FUNCTION "FC1041_TT_Taktimpuls" : Void   // FC1041, STL
TITLE = Taktimpuls bilden
{ S7_Optimized_Access := 'FALSE' }
AUTHOR : KT242
VERSION : 0.1
   VAR_INPUT
      IN_Drehfreigabe : Bool;   // Allgemeine Freigabe zum ansteuern der Anlage
      IN_Taktfreigabe : Bool;   // Freigabe zum Weitertakten der Anlage
      IN_Anlage_in_Position : Bool;   // Die Anlage befindet sich in der vorgegebenen Position
      IN_Start_Anlagenbetrieb : Bool;   // Die Anlage befindet sich in der Vorbereitung zum Produktionsbetrieb
      IN_Anlagenbetrieb : Bool;   // Die Anlage befindet sich im Produktionsbetrieb
      IN_DW_Taktzeit : S5Time;   // Zeitwert für die Taktzeit (Lauf- und Pausenzeit) der Anlage
      IN_Takttimer : Timer;   // Timer für die Bildung des Taktimpulses
      IN_Vorwarnzeit_1_in_Dec : Int;   // Zeitwert in Sekunden für eine Anfahrwarnung 1 vor dem Weitertakten
      IN_Vorwarnzeit_2_in_Dec : Int;   // Zeitwert in Sekunden für eine Anfahrwarnung 2 vor dem Weitertakten
   END_VAR
   VAR_IN_OUT
      IO_Status : "UDT_RT_Takt";   // Speichern der Takt- Zustände für das Programm
   END_VAR
   VAR_TEMP
      Temp_Restzeit : Int;   // Hilfwort mit Restzeit der Taktzeit in Sekunden
      Temp_Zeitraster : Byte;   // Hilfsbyte für dei ermittlung des Zeitrasters für die Bildung der Vorwarnungen
   END_VAR
BEGIN

REGION Network 1: Baustein abloeschen, wenn nicht Automatik
         O     #IN_Anlagenbetrieb;
         O     #IN_Start_Anlagenbetrieb;
         JC    NW1e;
   //
         R     #IO_Status.Vorwarnung_1;
         R     #IO_Status.Vorwarnung_2;
         R     #IO_Status.Taktzeit_beendet;
         R     #IO_Status.Taktimpuls;
         CLR;
         L     S5T#0MS;
         SP    #IN_Takttimer;
         BE;
   //
   NW1e: NOP   0;
END_REGION

REGION Network 2: Taktimpuls bilden
         L     #IN_DW_Taktzeit;
         A     #IN_Taktfreigabe;
         A     #IN_Drehfreigabe;
         A     #IO_Status.Taktzeit_beendet;
         SE    #IN_Takttimer;
         =     #IO_Status.Taktimpuls;
   //
         AN    #IN_Takttimer;
         =     #IO_Status.Taktzeit_beendet;
END_REGION

REGION Network 3: Vorwarnungsbits
   // Die Vorwarnungen werden nur gebildet, wenn sowohl bei der Taktzeit, als auch
   // bei den Vorwarnzeiten ein Sekundenzeitraster gewaehlt wurde
         LC    #IN_Takttimer;
         SRW   12;  // Zeitraster ermitteln
         T     #Temp_Zeitraster;
   //
         L     #Temp_Zeitraster;
         JL    wrne;
         JU    rst0;
         JU    rst1;
         JU    rst2;
         JU    rst3;
   wrne: JU    res;
   //
   rst0: L     #IN_Takttimer;
         L     100;
         /I;
         T     #Temp_Restzeit;
         JU    WRN;
   rst1: L     #IN_Takttimer;
         L     10;
         /I;
         T     #Temp_Restzeit;
         JU    WRN;
   rst2: L     #IN_Takttimer;
         L     1;
         /I;
         T     #Temp_Restzeit;
         JU    WRN;
   rst3: L     #IN_Takttimer;
         L     10;
         *I;
         T     #Temp_Restzeit;
         JU    WRN;
   //
   WRN:  L     #Temp_Restzeit;
         L     #IN_Vorwarnzeit_1_in_Dec;
         <I;
         =     #IO_Status.Vorwarnung_1;
         L     #Temp_Restzeit;
         L     #IN_Vorwarnzeit_2_in_Dec;
         <I;
         =     #IO_Status.Vorwarnung_2;
   //
         JU    nwe;
   res:  R     #IO_Status.Vorwarnung_1;
         R     #IO_Status.Vorwarnung_2;
   nwe:  NOP   0;
END_REGION
END_FUNCTION

FUNCTION "FC1042_RT_IPOS_CTRL" : Void   // FC1042, STL
TITLE = IPOS ansteuern
{ S7_Optimized_Access := 'FALSE' }
AUTHOR : KT242
VERSION : 0.1
// NEU 14.1.: Nach Quitt AS dreht RT ohne Warnung das Segment zu Ende
// NEU 23.1.: Start an FU wird jetzt gesetzt, auch wenn Umrichter nicht 
// betriebsbereit meldet. Es wird eine STG angezeigt und das Startbit wird mit 
// auslösen der STG reset. Somit erhält der Bediener eine Info, daß FU nicht 
// bereit 
// ist.
   VAR_INPUT
      IN_EA_Adresse : Hw_Any;   // Erste Adresse der Eingänge vom/ Ausgänge an den Umrichter
      IN_Taktend : Bool;   // Handelt es sich um einen taktenden Rundtisch?
      IN_Taktend_1_Segment : Bool;   // Soll im Automatikbetrieb durch Tippen positiv 1 Segment getaktet werden?
      IN_DP_ok : Bool;   // Ist der Umrichter am Profibus- System der Anlage erreichbar
      IN_IPOS_referenziert : Bool;   // Eingang das der Umrichter referenziert wurde
      IN_Stoerung_Luefter : Bool;   // Eingang Störung der Versorgung oder des Motorschutzes des Lüfters
      IN_Motorschutz : Bool;   // Eingang Störung der Versorgung oder des Motorschutzes des Umrichters
      IN_STG_Umrichter : Bool;   // Eingang Störung vom Frequenzumrichter
      IN_Reset_fault_Fkt : Bool;   // Signal zum quittieren der Störungen innerhalb der einzelnen Funktionsbausteine
      IN_Kettenspanner_ok : Bool;   // Signal vom Kettenspanner, Kette ist in Ordnung
      IN_Drehsperre : Bool;   // Es ist eine absolute Drehsperre eingeschaltet
      IN_HW_und_BA_ok : Bool;   // Eine gültige Betriebsart wurde angewählt und Steuerspannung ist aktiv
      IN_AutoStop_ok : Bool;   // Autostop ist ok bzw. quittiert
      IN_BA_Hand : Bool;   // Die Anlage befindet sich im Hand- Betrieb
      IN_BA_Automatik : Bool;   // Die Anlage befindet sich im Automatik- Betrieb
      IN_BA_Referenzieren : Bool;   // Die Anlage befindet sich im Referenzier- Betrieb
      IN_BA_Start_Taktbetrieb : Bool;   // Die Anlage befindet sich in der Startvorbereitung zum Produktions- Betrieb
      IN_BA_Taktbetrieb : Bool;   // Die Anlage befindet sich im Produktions- Betrieb
      IN_BA_Stop_angefordert : Bool;   // Die Anlage soll in einer definierten Position gestoppt werden
      IN_BA_Lampentest : Bool;   // Es sollen die Anzeigen der Anlage auf Funktion getestet werden
      IN_Taktimpuls : Bool;   // Bei einer taktenden Anlage soll die nächste Position angefahren werden
      IN_T_Tippen_plus : Bool;   // Eingang für den Taster zum ansteuern der Anlage in positive Richtung
      IN_T_Tippen_minus : Bool;   // Eingang für den Taster zum ansteuern der Anlage in negative Richtung
      IN_Genauhaltini : Bool;   // Eingang für einen Genauhaltinitiator für die Überprüfung der Positionierung
      IN_Anzahl_Segmente : Int;   // Anzahl der Segmente die sich innerhalb der 360° befinden
      IN_DW_Rampe_Pos : Int;   // Wert für die Beschleunigungsrampe des Umrichters (in ms)
      IN_DW_Rampe_Neg : Int;   // Wert für die Verzögerungssrampe des Umrichters (in ms)
      IN_DW_Speed_Hand : Int;   // Wert für die maximale Geschwindigkeit in der Betriebsart Tippen Hand
      IN_DW_Speed_Automatik : Int;   // Wert für die maximale Geschwindigkeit in der Betriebsart Automatik
      IN_DW_Offset_Position : Int;   // Wert des "negativen" Offset der Positionierung bei kontinuierlichem Rundtisch
      IN_TM_Universal : Timer;   // Timer für die Betriebsart und die Taktverzögerung des Rundtisches
      IN_TM_Freigabe : Timer;   // Timer für die Ausschaltverzögerung der Umrichterfreigaben
      IN_TM_Tol_Genauhalt : Timer;   // Timer für die Überwachung der Genauhaltepositin
      IN_TM_Verz_STG_FU : Timer;   // Timer für Verzögerung Stg FU
      IN_TM_Verz_Ziel_erreicht : Timer;
      IN_TM_AnfahrWarnung : Timer;   // Timer für die Ausgabe einer Anfahrwarnung
      IN_ZT_Tol_Genauhalt : S5Time;   // Zeitwert für die Überwachung der Genauhalteposition
      IN_Time_Anfahrwarnung : S5Time;   // Zeitwert für die Anfahrwarnung
   END_VAR
   VAR_OUTPUT
      OUT_aktuelle_Position : Int;   // Wert mit der aktuellen Position innerhalb des Segmentes (in 1/10 Grad)
      OUT_FRG_Umrichter : Bool;   // Ausgang für die Hardware- Freigabe des Umrichters
      OUT_H_Tippen_plus : Bool;   // Ausgang für die Anzeige Tippen positiv
      OUT_H_Tippen_minus : Bool;   // Ausgang für die Anzeige Tippen negativ
      OUT_H_Referenzpunkt : Bool;   // Ausgang für die Anzeige der Referenzierung
      OUT_H_AnfahrWarnung : Bool;   // Ausgang für die ANsteuerung der ANfahrwarnung
   END_VAR
   VAR_IN_OUT
      IO_Status : "UDT_RT_IPOS";   // Speichern des Umrichter- Status und der Ein- und Ausgänge für das Programm
      IO_Fault : Struct
         STG_Luefter : Bool;   // Störung: Der Versorgung oder des Motorschutzes des Lüfters
         STG_Umrichter : Bool;   // Störung: Der Umrichter ist nicht betriebsbereit
         STG_Motorschutz : Bool;   // Störung: Der Versorgung oder des Motorschutzes des Umrichters
         STG_von_IPOS : Bool;   // Störung: Ein Störungssignal von dem Umrichter steht an
         STG_Genauhaltini : Bool;   // Störung: Die Genauhalteposition (Initiator) wurde nicht erreicht
         STG_Genauhalt_immer_ein : Bool;   // Störung: Die Genauhalteposition (Initiator) wird dauernd belegt
         STG_Busfehler : Bool;   // Störung: Busteilnehmer ist nicht erreichbar
         STG_Reserve_0_7 : Bool;
         STG_Reserve_1_0 : Bool;
         STG_Reserve_1_1 : Bool;
         STG_Reserve_1_2 : Bool;
         STG_Reserve_1_3 : Bool;
         STG_Reserve_1_4 : Bool;
         STG_Reserve_1_5 : Bool;
         STG_Reserve_1_6 : Bool;
         STG_Reserve_1_7 : Bool;
      END_STRUCT;
      IO_New_Fault : Bool;   // Eine neue Störung steht an
      IO_Fault_GRP_1 : Bool;   // Eine Störungd er Gruppe 1 steht an
      IO_Fault_GRP_2 : Bool;   // Eine Störungd er Gruppe 2 steht an
      IO_Fault_GRP_3 : Bool;   // Eine Störungd er Gruppe 3 steht an
   END_VAR
   VAR_TEMP
      Temp_IO_Status : "UDT_RT_IPOS";   // Temporärer Umrichter- Status für die interne Bearbeitung des Bausteins
      ERROR_CODE : Int;   // Störungszustand der Systemfunktion "BLKMOV" Blockmove
      Anyzeiger : ANY;   // Zeiger zum Kopieren der Bereiche "IO_Status" und "Temp_IO_Status"
      Temp_Nullmerker : Int;   // Nullmerker zum ablöschen der Eingänge bei Profibus- Störungen
      Temp_Segmentbreite : DInt;   // Die breite eines Segmentes in 1/10 Grad (Summe aller Segmente = 3600)
      Temp_aktuelle_Position : DInt;   // Die aktuelle Position innerhalb eines Segmentes
      Temp_BA_Wechsel : Bool;   // Hilfsmerker: Es wurde ein wechsel der Betriebsart festgestellt
      Temp_BA_Time : Bool;   // Hilfsmerker: Die Wartezeit zur Erkennung der Betriebsart ist abgelaufen
      Temp_FRG_Bewegung : Bool;   // Hilfsmerker: Eine Ansteuerung des Umrichters ist Freigegeben
      Temp_FIM_BA_Referenz : Bool;   // Hilfsmerker: Flankenimpuls zum Starten des Referenzierens der Anlage
      Temp_FIM_Referenz : Bool;   // Hilfsmerker: Flankenimpuls für die Erkennung der Genauhalteposition
      Temp_FIM_Tip_Auto : Bool;   // Hilfsmerker: Flankenimpuls für das Weitertakten im automatischen Tip- Betrieb
      Temp_neues_Ziel : Bool;   // Hilfsmerker: Freigabe zum berechnen eines neuen Zieles bei kontinuierlichen RT
      Temp_Freigabe_Stopp : Bool;   // Hilfsmerker: Freigabe zum Stoppen des Rundtisches
   END_VAR
BEGIN

REGION Network 1: Gesicherte Daten einbinden
         LAR1;
         L;
         LAR2;
   //
         L     W#16#1002;  // Bytes
         T     W[AR1, P#0.0];
         L     40;  // Anzahl Bytes
         T     W[AR1, P#2.0];
         L     W[AR2, P#0.0];  // Baustein Nr.
         T     W[AR1, P#4.0];
         L     D[AR2, P#2.0];  // Datenanfang
         T     D[AR1, P#6.0];
   //
         CALL  BLKMOV
         ( SRCBLK  := #Anyzeiger,
           RET_VAL := #ERROR_CODE,
           DSTBLK  := #Temp_IO_Status
         );
   //
END_REGION

REGION Network 2: Anstehende Störungen zurücksetzen
   //-----
         A     #IN_Reset_fault_Fkt;
         R     #IO_Fault.STG_Luefter;
         R     #IO_Fault.STG_Umrichter;
         R     #IO_Fault.STG_Motorschutz;
         R     #IO_Fault.STG_von_IPOS;
         R     #IO_Fault.STG_Genauhaltini;
         R     #IO_Fault.STG_Genauhalt_immer_ein;
         R     #IO_Fault.STG_Busfehler;
   //-----
END_REGION

REGION Network 3: Eingänge von IPOS laden
   // Um ein permanentes Beschreiben des Diagnosepuffers zu verhindern, werden die 
   // Peripheriebefehle übersprungen, sobald festgestellt wurde, daß der Teilnehmer 
   // ausgefallen ist.
         L     0;
         T     #Temp_Nullmerker;
   //
         AN    #IN_DP_ok;
         JC    pae0;
   //
         CALL  DPRD_DAT
         ( LADDR   := #IN_EA_Adresse,
           RET_VAL := #ERROR_CODE,
           RECORD  := #Temp_IO_Status.Eingaenge_von_IPOS
         );
   //
         JU    paee;
   pae0: NOP   0;
   //-
         AN    #IN_DP_ok;
         AN    #IO_Fault.STG_Busfehler;
         S     #IO_Fault.STG_Busfehler;
         S     #IO_New_Fault;
   //-
         CALL  FILL
         ( BVAL    := #Temp_Nullmerker,
           RET_VAL := #ERROR_CODE,
           BLK     := #Temp_IO_Status.Eingaenge_von_IPOS
         );
   //
   paee: NOP   0;
   //
END_REGION

REGION Network 4: aktuelle Position
         L     3600;  // 360° Umfang
         L     #IN_Anzahl_Segmente;  // Anzahl der Segmente
         /D;
         T     #Temp_Segmentbreite;  // in 1/10 Grad
   //__________________________________________________________________
   //
         L     #Temp_IO_Status.Eingaenge_von_IPOS.Istposition;
         L     #Temp_Segmentbreite;  // in 1/10 Grad
         MOD;
         T     #Temp_aktuelle_Position;  // Aktuelle Position im Segment
         T     #Temp_IO_Status.Status.Aktuelle_Position;
         T     #OUT_aktuelle_Position;
END_REGION

REGION Network 5: Position erreicht
   // Zeil erreicht nur zulassen wenn auf 0 Teilung
         L     #Temp_IO_Status.Status.Aktuelle_Position;
         L     0;
         ==I;
         A     #Temp_IO_Status.Eingaenge_von_IPOS.Ziel_erreicht;
         =     #Temp_IO_Status.Eingaenge_von_IPOS.Ziel_erreicht;
END_REGION

REGION Network 6: Störungsauswertung
         A     #Temp_IO_Status.Eingaenge_von_IPOS.Stoerung_Warnung;
         A     #IN_Reset_fault_Fkt;
         =     #Temp_IO_Status.Ausgaenge_an_IPOS.Reset;
   //
         A     #IN_Stoerung_Luefter;
         AN    #IO_Fault.STG_Luefter;
         S     #IO_Fault.STG_Luefter;
         S     #IO_New_Fault;
         S     #IO_Fault_GRP_3;
   //
   //----NEU 23.1.
         A     #Temp_IO_Status.Ausgaenge_an_IPOS.DI_00_Start;
         O     #Temp_IO_Status.Ausgaenge_an_IPOS.DI_01_T_plus;
         O     #Temp_IO_Status.Ausgaenge_an_IPOS.DI_02_T_minus;
         AN    #Temp_IO_Status.Eingaenge_von_IPOS.Umrichter_betriebsbereit;
         L     S5T#1S_500MS;
         SD    #IN_TM_Verz_STG_FU;
         A     #IN_TM_Verz_STG_FU;
         AN    #IO_Fault.STG_Umrichter;
         S     #IO_Fault.STG_Umrichter;
         S     #IO_New_Fault;
         S     #IO_Fault_GRP_1;
   //-----
         O     #Temp_IO_Status.Eingaenge_von_IPOS.Stoerung_Warnung;
         ON    #IN_STG_Umrichter;
         AN    #Temp_IO_Status.Ausgaenge_an_IPOS.Reset;
         AN    #IO_Fault.STG_von_IPOS;
         S     #IO_Fault.STG_von_IPOS;
         S     #IO_New_Fault;
         S     #IO_Fault_GRP_3;
   //
         A     #IN_Motorschutz;
         AN    #IO_Fault.STG_Motorschutz;
         S     #IO_Fault.STG_Motorschutz;
         S     #IO_New_Fault;
         S     #IO_Fault_GRP_1;
   //-----
         A(;
         L     #Temp_Segmentbreite;
         L     10;
         *D;
         L     100;
         /D;
         L     #Temp_aktuelle_Position;
         <D;
         );
         AN(;
         L     #Temp_Segmentbreite;
         L     90;
         *D;
         L     100;
         /D;
         L     #Temp_aktuelle_Position;
         <D;
         );
         O     #Temp_IO_Status.Status.BA_Referenzieren;
         ON    #Temp_IO_Status.Status.IPOS_referenziert;
         R     #Temp_IO_Status.Status.HM_Chk_Genauhalt_ok;
   //
         AN(;
         A     #IN_BA_Hand;
         A     #Temp_IO_Status.Status.BA_Tippen;
         );
         A(;
         L     #Temp_Segmentbreite;
         L     98;
         *D;
         L     100;
         /D;
         L     #Temp_aktuelle_Position;
         <D;
         );
         AN    #Temp_IO_Status.Status.HM_Chk_Genauhalt_ok;
         FP    #Temp_IO_Status.Status.FHM_STG_Genauhaltini;
         S     #Temp_IO_Status.Status.HM_STG_Chk_Genauhalt;
   //
         O     #IN_Genauhaltini;
         O     #IO_Fault.STG_Genauhaltini;
         A     #Temp_IO_Status.Status.HM_STG_Chk_Genauhalt;
         R     #Temp_IO_Status.Status.HM_STG_Chk_Genauhalt;
         S     #Temp_IO_Status.Status.HM_Chk_Genauhalt_ok;
         S     #IO_Fault_GRP_1;
   //
         A     #IN_Taktend;
         A     #Temp_IO_Status.Eingaenge_von_IPOS.Ziel_erreicht;
         AN    #IN_Genauhaltini;
         O;
         AN    #IN_Taktend;
         AN    #IN_BA_Stop_angefordert;
         AN    #Temp_IO_Status.Status.BA_Referenzieren;
         A     #Temp_IO_Status.Status.HM_STG_Chk_Genauhalt;
         L     #IN_ZT_Tol_Genauhalt;
         SD    #IN_TM_Tol_Genauhalt;
         A     #IN_TM_Tol_Genauhalt;
         AN    #IO_Fault.STG_Genauhaltini;
         S     #IO_Fault.STG_Genauhaltini;
         S     #IO_New_Fault;
         S     #IO_Fault_GRP_1;
   //
         A     #Temp_IO_Status.Ausgaenge_an_IPOS.DI_00_Start;
         FP    #Temp_IO_Status.Status.FHM_STG_Start;
         R     #Temp_IO_Status.Status.Genauhalt_war_verlassen;
         ON    #IN_Genauhaltini;
         S     #Temp_IO_Status.Status.Genauhalt_war_verlassen;
   //
         A     #Temp_IO_Status.Status.RT_in_Position;
         FP    #Temp_IO_Status.Status.FHM_STG_in_Position;
         A     #IN_Genauhaltini;
         AN    #Temp_IO_Status.Ausgaenge_an_IPOS.DI_00_Start;
         AN    #Temp_IO_Status.Status.Genauhalt_war_verlassen;
         AN    #IO_Fault.STG_Genauhalt_immer_ein;
         S     #IO_Fault.STG_Genauhalt_immer_ein;
         S     #IO_New_Fault;
         S     #IO_Fault_GRP_1;
   //-----
END_REGION

REGION Network 7: Betriebsarten anwählen
         CLR;
         =     #Temp_BA_Wechsel;
   //
         A     #IN_BA_Hand;
         A     #IN_BA_Referenzieren;
         JC    BA_r;
         O     #IN_BA_Start_Taktbetrieb;
         O     #IN_BA_Taktbetrieb;
         O;
         A     #IN_Taktend_1_Segment;
         A     #IN_BA_Automatik;
         AN    #IN_BA_Start_Taktbetrieb;
         AN    #IN_BA_Taktbetrieb;
         JC    BA_a;
         AN    #IN_BA_Hand;
   //    UN    #IN_BA_Automatik
         JC    BA_c;
   //___________________________________________________________
   // Betriebsart Tippbetrieb
         ON    #Temp_IO_Status.Ausgaenge_an_IPOS.DI_03_Mode_Tipp;
         O     #Temp_IO_Status.Ausgaenge_an_IPOS.DI_04_Mode_Ref;
         O     #Temp_IO_Status.Ausgaenge_an_IPOS.DI_05_Mode_Auto;
         =     #Temp_BA_Wechsel;
         SET;
         S     #Temp_IO_Status.Ausgaenge_an_IPOS.DI_03_Mode_Tipp;
         R     #Temp_IO_Status.Ausgaenge_an_IPOS.DI_04_Mode_Ref;
         R     #Temp_IO_Status.Ausgaenge_an_IPOS.DI_05_Mode_Auto;
         JU    BA_e;
   //___________________________________________________________
   // Betriebsart Referenzieren
   BA_r: O     #Temp_IO_Status.Ausgaenge_an_IPOS.DI_03_Mode_Tipp;
         ON    #Temp_IO_Status.Ausgaenge_an_IPOS.DI_04_Mode_Ref;
         O     #Temp_IO_Status.Ausgaenge_an_IPOS.DI_05_Mode_Auto;
         =     #Temp_BA_Wechsel;
         SET;
         R     #Temp_IO_Status.Ausgaenge_an_IPOS.DI_03_Mode_Tipp;
         S     #Temp_IO_Status.Ausgaenge_an_IPOS.DI_04_Mode_Ref;
         R     #Temp_IO_Status.Ausgaenge_an_IPOS.DI_05_Mode_Auto;
         JU    BA_e;
   //___________________________________________________________
   // Betriebsart Automatik
   BA_a: O     #Temp_IO_Status.Ausgaenge_an_IPOS.DI_03_Mode_Tipp;
         O     #Temp_IO_Status.Ausgaenge_an_IPOS.DI_04_Mode_Ref;
         ON    #Temp_IO_Status.Ausgaenge_an_IPOS.DI_05_Mode_Auto;
         =     #Temp_BA_Wechsel;
         SET;
         R     #Temp_IO_Status.Ausgaenge_an_IPOS.DI_03_Mode_Tipp;
         R     #Temp_IO_Status.Ausgaenge_an_IPOS.DI_04_Mode_Ref;
         S     #Temp_IO_Status.Ausgaenge_an_IPOS.DI_05_Mode_Auto;
         JU    BA_e;
   //___________________________________________________________
   // Betriebsarten ablöschen
   BA_c: O     #Temp_IO_Status.Ausgaenge_an_IPOS.DI_03_Mode_Tipp;
         O     #Temp_IO_Status.Ausgaenge_an_IPOS.DI_04_Mode_Ref;
         O     #Temp_IO_Status.Ausgaenge_an_IPOS.DI_05_Mode_Auto;
         =     #Temp_BA_Wechsel;
         SET;
         R     #Temp_IO_Status.Ausgaenge_an_IPOS.DI_03_Mode_Tipp;
         R     #Temp_IO_Status.Ausgaenge_an_IPOS.DI_04_Mode_Ref;
         R     #Temp_IO_Status.Ausgaenge_an_IPOS.DI_05_Mode_Auto;
         JU    BA_e;
   BA_e: NOP   0;
END_REGION

REGION Network 8: Wartezeit zwischen Betriebsart und Ansteuerung
         AN    #Temp_BA_Wechsel;
         JC    Ba_T;
   //
         CLR;
         L     S5T#0MS;
         SP    #IN_TM_Universal;
         SET;
         R     #Temp_IO_Status.Status.BA_Tippen;
         R     #Temp_IO_Status.Status.BA_Referenzieren;
         R     #Temp_IO_Status.Status.BA_Takt_Automatik;
         R     #Temp_IO_Status.Status.BA_Produktion;
         R     #Temp_IO_Status.Status.BA_Produktion_Kont;
         R     #Temp_IO_Status.Status.BA_gueltig;
         JU    Ba_Eä;
   //
   Ba_T: NOP   0;
   //
         A     #Temp_IO_Status.Status.BA_gueltig;
         JC    Ba_Eä;
   //
         O     #Temp_IO_Status.Ausgaenge_an_IPOS.DI_03_Mode_Tipp;
         O     #Temp_IO_Status.Ausgaenge_an_IPOS.DI_04_Mode_Ref;
         O     #Temp_IO_Status.Ausgaenge_an_IPOS.DI_05_Mode_Auto;
         AN    #Temp_BA_Wechsel;
         L     S5T#250MS;
         SD    #IN_TM_Universal;
   //
         A     #IN_TM_Universal;
         =     #Temp_BA_Time;
         S     #Temp_IO_Status.Status.BA_gueltig;
   //
         A     #Temp_BA_Time;
         A     #IN_BA_Hand;
         A     #Temp_IO_Status.Ausgaenge_an_IPOS.DI_03_Mode_Tipp;
         S     #Temp_IO_Status.Status.BA_Tippen;
   //
         A     #Temp_BA_Time;
         A     #IN_BA_Automatik;
         AN    #IN_Taktend_1_Segment;
         A     #Temp_IO_Status.Ausgaenge_an_IPOS.DI_03_Mode_Tipp;
         S     #Temp_IO_Status.Status.BA_Tippen;
   //
         A     #Temp_BA_Time;
         A     #Temp_IO_Status.Ausgaenge_an_IPOS.DI_04_Mode_Ref;
         S     #Temp_IO_Status.Status.BA_Referenzieren;
   //
         A     #Temp_BA_Time;
         A     #IN_Taktend_1_Segment;
         A     #IN_Taktend;
         A     #Temp_IO_Status.Ausgaenge_an_IPOS.DI_05_Mode_Auto;
         S     #Temp_IO_Status.Status.BA_Takt_Automatik;
   //
         A     #Temp_BA_Time;
         A     #IN_Taktend;
         A     #Temp_IO_Status.Ausgaenge_an_IPOS.DI_05_Mode_Auto;
         S     #Temp_IO_Status.Status.BA_Produktion;
   //
         A     #Temp_BA_Time;
         AN    #IN_Taktend;
         A     #Temp_IO_Status.Ausgaenge_an_IPOS.DI_05_Mode_Auto;
         S     #Temp_IO_Status.Status.BA_Produktion_Kont;
   //
         AN    #Temp_IO_Status.Status.BA_gueltig;
         JC    Ba_Eä;
   //
         CLR;
         L     S5T#0MS;
         SP    #IN_TM_Universal;
   //
   Ba_Eä:NOP   0;
END_REGION

REGION Network 9: Funktionsbits ablöschen bei Betriebsartenwechsel
         ON    #Temp_IO_Status.Status.BA_gueltig;
         ON    #IN_AutoStop_ok;
         O     #IO_Fault.STG_Umrichter;
         R     #Temp_IO_Status.Ausgaenge_an_IPOS.DI_00_Start;
         R     #Temp_IO_Status.Ausgaenge_an_IPOS.DI_01_T_plus;
         R     #Temp_IO_Status.Ausgaenge_an_IPOS.DI_02_T_minus;
         R     #Temp_IO_Status.Status.RT_dreht;
         R     #Temp_IO_Status.Status.Stoppen_erkannt;
END_REGION

REGION Network 10: Bewegungen freigeben
   // NEU 23.1.:Umrichter_betriebsbereit raus, damit DI_00_Start gesetzt werden kann 
   // im NW13
         AN    #IO_Fault.STG_Umrichter;
         AN    #IO_Fault.STG_Motorschutz;
         AN    #IO_Fault.STG_von_IPOS;
         A     #Temp_IO_Status.Status.BA_gueltig;
         A     #IN_HW_und_BA_ok;
         A     #IN_Kettenspanner_ok;
         AN    #IN_Drehsperre;
         A     #IN_AutoStop_ok;
         =     #Temp_FRG_Bewegung;
END_REGION

REGION Network 11: Tippbetrieb Hand
         A     #IN_BA_Hand;
         A     #Temp_IO_Status.Status.BA_Tippen;
         JCN   etpH;
   //
         A     #IN_T_Tippen_plus;
         AN    #IN_T_Tippen_minus;
         A     #Temp_FRG_Bewegung;
         =     #Temp_IO_Status.Ausgaenge_an_IPOS.DI_01_T_plus;
   //
         AN    #IN_T_Tippen_plus;
         A     #IN_T_Tippen_minus;
         A     #Temp_FRG_Bewegung;
         =     #Temp_IO_Status.Ausgaenge_an_IPOS.DI_02_T_minus;
   //
         O     #Temp_IO_Status.Ausgaenge_an_IPOS.DI_01_T_plus;
         O     #Temp_IO_Status.Ausgaenge_an_IPOS.DI_02_T_minus;
         R     #Temp_IO_Status.Status.RT_in_Position;
         R     #Temp_IO_Status.Status.Ziel_ermittelt;
   //
         L     #IN_DW_Speed_Hand;
         T     #Temp_IO_Status.Status.Ziel_Geschwindigkeit;
   //
         L     #IN_DW_Rampe_Pos;
         T     #Temp_IO_Status.Status.Ziel_Beschleunigung;
   //
         L     #IN_DW_Rampe_Neg;
         T     #Temp_IO_Status.Status.Ziel_Verzoegerung;
   //
   etpH: NOP   0;
END_REGION

REGION Network 12: Tippbetrieb Automatik
         A     #IN_BA_Automatik;
         A     #Temp_IO_Status.Status.BA_Tippen;
         JCN   etpA;
   //
         A     #IN_T_Tippen_plus;
         AN    #IN_T_Tippen_minus;
         A     #Temp_FRG_Bewegung;
         =     #Temp_IO_Status.Ausgaenge_an_IPOS.DI_01_T_plus;
   //
         A     #Temp_IO_Status.Ausgaenge_an_IPOS.DI_01_T_plus;
         R     #Temp_IO_Status.Status.RT_in_Position;
         R     #Temp_IO_Status.Status.Ziel_ermittelt;
   //
         L     #IN_DW_Speed_Automatik;
         T     #Temp_IO_Status.Status.Ziel_Geschwindigkeit;
   //
         L     #IN_DW_Rampe_Pos;
         T     #Temp_IO_Status.Status.Ziel_Beschleunigung;
   //
         L     #IN_DW_Rampe_Neg;
         T     #Temp_IO_Status.Status.Ziel_Verzoegerung;
   //
   etpA: NOP   0;
END_REGION

REGION Network 13: Referenzieren
         A     #Temp_IO_Status.Status.BA_Referenzieren;
         FP    #Temp_IO_Status.Status.FHM_BA_Referenzieren;
         =     #Temp_FIM_BA_Referenz;
   //
         A     #IN_BA_Hand;
         A     #IN_BA_Referenzieren;
         A     #Temp_IO_Status.Status.BA_Referenzieren;
         JCN   eref;
   //
         A     #Temp_FIM_BA_Referenz;
         R     #Temp_IO_Status.Status.RT_in_Position;
         R     #Temp_IO_Status.Status.Ziel_ermittelt;
   //
         A     #Temp_FIM_BA_Referenz;
         S     #Temp_IO_Status.Ausgaenge_an_IPOS.DI_00_Start;
   //
         A     #IN_IPOS_referenziert;
         FP    #Temp_IO_Status.Status.FHM_Referenziert;
         =     #Temp_FIM_Referenz;
   //
         A     #Temp_FIM_Referenz;
         A     #IN_Genauhaltini;
         S     #Temp_IO_Status.Status.RT_in_Position;
   //
         A     #Temp_FIM_Referenz;
         R     #Temp_IO_Status.Ausgaenge_an_IPOS.DI_00_Start;
         JCN   tghl;
         L     0;
         T     #Temp_IO_Status.Status.Ziel_Position;
   //
   tghl: A     #Temp_FIM_Referenz;
         AN    #IN_Genauhaltini;
         AN    #IO_Fault.STG_Genauhaltini;
         S     #IO_Fault.STG_Genauhaltini;
         S     #IO_Fault_GRP_1;
   eref: NOP   0;
END_REGION

REGION Network 14: Automatik // Tip- Betrieb
         A     #Temp_IO_Status.Status.BA_Takt_Automatik;
         JCN   ea_T;
   //
         A     #IN_T_Tippen_plus;
         AN    #IN_T_Tippen_minus;
         AN    #Temp_IO_Status.Status.RT_dreht;
         AN    #IN_BA_Stop_angefordert;
         FP    #Temp_IO_Status.Status.FHM_Auto_kont;
         =     #Temp_FIM_Tip_Auto;
   //___________________________________________________________________________
   // Ziel für Bewegung ermitteln
         AN    #Temp_IO_Status.Status.RT_dreht;
         AN    #Temp_IO_Status.Status.Ziel_ermittelt;
         AN    #Temp_IO_Status.Ausgaenge_an_IPOS.DI_00_Start;
         JCN   T_aT;
         S     #Temp_IO_Status.Status.Ziel_ermittelt;
   //
         A     #Temp_IO_Status.Status.RT_in_Position;
         AN(;
         L     #Temp_IO_Status.Eingaenge_von_IPOS.Istposition;
         L     #Temp_IO_Status.Status.Ziel_Position;
         ==D;
         );
         JC    G_at;
   // Start aus Zwischenposition
         L     #Temp_IO_Status.Eingaenge_von_IPOS.Istposition;
         L     #Temp_aktuelle_Position;
         -D;
         L     #Temp_Segmentbreite;
         +D;
         T     #Temp_IO_Status.Status.Ziel_Position;
         JU    T_aT;
   //
   // Start aus Genauhaltposition
   G_at: L     #Temp_IO_Status.Status.Ziel_Position;
         L     #Temp_Segmentbreite;
         +D;
         L     3600;  // 360° Umfang
         MOD;
         T     #Temp_IO_Status.Status.Ziel_Position;
   //___________________________________________________________________________
   // Rundtisch weiter takten
   T_aT: NOP   0;
         A     #Temp_FIM_Tip_Auto;
         JCN   bewT;
         S     #Temp_IO_Status.Status.RT_dreht;
         R     #Temp_IO_Status.Status.RT_in_Position;
         R     #Temp_IO_Status.Status.Ziel_ermittelt;
   //
   // Bewegung starten und Steuersignale ausgeben
   bewT: NOP   0;
   //
         A     #IN_Genauhaltini;
         A     #Temp_IO_Status.Eingaenge_von_IPOS.Ziel_erreicht;
         FP    #Temp_IO_Status.Status.FHM_RT_in_Position;
         R     #Temp_IO_Status.Status.RT_dreht;
         S     #Temp_IO_Status.Status.RT_in_Position;
   //--------------------------
         L     #IN_DW_Speed_Automatik;
         T     #Temp_IO_Status.Status.Ziel_Geschwindigkeit;
   //--------------------------
         L     #IN_DW_Rampe_Pos;
         T     #Temp_IO_Status.Status.Ziel_Beschleunigung;
   //
         L     #IN_DW_Rampe_Neg;
         T     #Temp_IO_Status.Status.Ziel_Verzoegerung;
   //--------------------------
   // Nachlaufzeit für Positionierung
         A     #Temp_IO_Status.Status.RT_dreht;
         L     S5T#500MS;
         SF    #IN_TM_Universal;
         A     #IN_TM_Universal;
         A     #Temp_FRG_Bewegung;
         =     #Temp_IO_Status.Ausgaenge_an_IPOS.DI_00_Start;
   ea_T: NOP   0;
END_REGION

REGION Network 15: Automatik // Taktbetrieb
         O     #IN_BA_Start_Taktbetrieb;
         O     #IN_BA_Taktbetrieb;
         A     #Temp_IO_Status.Status.BA_Produktion;
         JCN   ea_P;
   //___________________________________________________________________________
   // Anwahl zum Stoppen des Rundtischen
   //
         A     #IN_BA_Stop_angefordert;
         S     #Temp_IO_Status.Status.Stoppen_erkannt;
   //___________________________________________________________________________
   // Ziel für Bewegung ermitteln
   //
         AN    #Temp_IO_Status.Status.RT_dreht;
         AN    #Temp_IO_Status.Status.Ziel_ermittelt;
         AN    #Temp_IO_Status.Ausgaenge_an_IPOS.DI_00_Start;
         JCN   T_aP;
         S     #Temp_IO_Status.Status.Ziel_ermittelt;
   //
         A     #Temp_IO_Status.Status.RT_in_Position;
         JC    G_aP;
   // Start aus Zwischenposition
         L     #Temp_IO_Status.Eingaenge_von_IPOS.Istposition;
         L     #Temp_aktuelle_Position;
         -D;
         L     #Temp_Segmentbreite;
         +D;
         T     #Temp_IO_Status.Status.Ziel_Position;
         JU    T_aP;
   //
   // Start aus Genauhaltposition
   G_aP: L     #Temp_IO_Status.Status.Ziel_Position;
         L     #Temp_Segmentbreite;
         +D;
         L     3600;  // 360° Umfang
         MOD;
         T     #Temp_IO_Status.Status.Ziel_Position;
   //___________________________________________________________________________
   // Rundtisch weiter takten
   T_aP: NOP   0;
         A     #IN_Taktimpuls;
         JCN   bewP;
         S     #Temp_IO_Status.Status.RT_dreht;
         R     #Temp_IO_Status.Status.RT_in_Position;
         R     #Temp_IO_Status.Status.Ziel_ermittelt;
   //
   // Bewegung starten und Steuersignale ausgeben
   bewP: NOP   0;
   //
         A     #Temp_IO_Status.Eingaenge_von_IPOS.Ziel_erreicht;
         A     #IN_Genauhaltini;
         FP    #Temp_IO_Status.Status.FHM_RT_in_Position;
         R     #Temp_IO_Status.Status.RT_dreht;
         S     #Temp_IO_Status.Status.RT_in_Position;
   //--------------------------
         L     #IN_DW_Speed_Automatik;
         T     #Temp_IO_Status.Status.Ziel_Geschwindigkeit;
   //--------------------------
         L     #IN_DW_Rampe_Pos;
         T     #Temp_IO_Status.Status.Ziel_Beschleunigung;
   //
         L     #IN_DW_Rampe_Neg;
         T     #Temp_IO_Status.Status.Ziel_Verzoegerung;
   //--------------------------
   // Nachlaufzeit für Positionierung
         A     #Temp_IO_Status.Status.RT_dreht;
         L     S5T#500MS;
         SF    #IN_TM_Universal;
         A     #IN_TM_Universal;
         A     #Temp_FRG_Bewegung;
         =     #Temp_IO_Status.Ausgaenge_an_IPOS.DI_00_Start;
   ea_P: NOP   0;
END_REGION

REGION Network 16: Automatik - kontinuierlich drehend
         O     #IN_BA_Start_Taktbetrieb;
         O     #IN_BA_Taktbetrieb;
         A     #Temp_IO_Status.Status.BA_Produktion_Kont;
         JCN   ea_k;
   //___________________________________________________________________________
   // Ziel für Bewegung ermitteln
   //
   // Neue Zielvorgabe bei erreichen von 85% des Segmentes:
   //
         A(;
         L     #Temp_Segmentbreite;
         L     50;
         *D;
         L     100;
         /D;
         L     #Temp_aktuelle_Position;
         <D;
         );
         =     #Temp_neues_Ziel;
   //
   // Die Freigabe zum Stoppen wird erst gegeben wen 10% des Segmentes vorbei sind:
   //
         A(;
         L     #Temp_Segmentbreite;
         L     10;
         *D;
         L     100;
         /D;
         L     #Temp_aktuelle_Position;
         <D;
         );
         =     #Temp_Freigabe_Stopp;
   //
   // Anwahl zum Stoppen des Rundtischen
   //
         A     #IN_BA_Stop_angefordert;
         AN    #Temp_neues_Ziel;
         A     #Temp_Freigabe_Stopp;
         S     #Temp_IO_Status.Status.Stoppen_erkannt;
         AN    #IN_BA_Stop_angefordert;
         R     #Temp_IO_Status.Status.Stoppen_erkannt;
   //
         A     #Temp_neues_Ziel;
         A     #Temp_IO_Status.Status.RT_dreht;
         AN    #Temp_IO_Status.Status.Ziel_ermittelt;
         AN    #Temp_IO_Status.Status.Stoppen_erkannt;
         O;
         AN    #Temp_IO_Status.Status.RT_dreht;
         AN    #Temp_IO_Status.Status.Ziel_ermittelt;
         AN    #Temp_IO_Status.Ausgaenge_an_IPOS.DI_00_Start;
         AN    #Temp_IO_Status.Status.Stoppen_erkannt;
         JCN   T_aK;
   //
         AN    #IN_BA_Stop_angefordert;
         S     #Temp_IO_Status.Status.Ziel_ermittelt;
   //
         A     #Temp_neues_Ziel;
         A     #Temp_IO_Status.Status.RT_dreht;
         O     #Temp_IO_Status.Status.RT_in_Position;
         JC    G_aK;
   // Start aus Zwischenposition:
   // Start außerhalb des Bereiches für die neue Positionsvorgabe:
         L     #Temp_IO_Status.Eingaenge_von_IPOS.Istposition;
         L     #Temp_aktuelle_Position;
         -D;
         L     #Temp_Segmentbreite;
         +D;
         L     #IN_DW_Offset_Position;
         -D;
         T     #Temp_IO_Status.Status.Ziel_Position;
   // Bei start innerhalb des Bereiches für die neue Positionsvorgabe
   // wird gleich auf das nächste Zil verwiesen:
         A     #Temp_neues_Ziel;
         JCN   T_aK;
   // Start aus definierter Position heraus:
   // Während des Betriebs:
   G_aK: NOP   0;
         L     #Temp_IO_Status.Status.Ziel_Position;
         L     #Temp_Segmentbreite;
         +D;
         L     #IN_DW_Offset_Position;
         -D;
         L     3600;  // 360° Umfang
         MOD;
         T     #Temp_IO_Status.Status.Ziel_Position;
   //___________________________________________________________________________
   // Rundtisch weiter takten
   T_aK: NOP   0;

   //      L     #Temp_aktuelle_Position
   //      L     10
   //      >I
   //    )
         ON    #IN_Genauhaltini;
         FP    #Temp_IO_Status.Status.FHM_Auto_kont;
         R     #Temp_IO_Status.Status.RT_in_Position;
   //
         ON    #Temp_IO_Status.Status.RT_dreht;
         S     #Temp_IO_Status.Status.RT_dreht;
   //
         AN    #Temp_neues_Ziel;
         A     #Temp_Freigabe_Stopp;
         R     #Temp_IO_Status.Status.Ziel_ermittelt;
   //
   // Bewegung starten und Steuersignale ausgeben
         NOP   0;
   //
   //    O(
   //      L     #Temp_Segmentbreite
   //      L     10
   //      *D
   //      L     100
   //      /D
   //      L     #Temp_aktuelle_Position
   //      <D
   //    )
         O     #IN_Genauhaltini;
         FP    #Temp_IO_Status.Status.FHM_RT_in_Position;
         S     #Temp_IO_Status.Status.RT_in_Position;
   //--------------------------
         L     #IN_DW_Speed_Automatik;
         T     #Temp_IO_Status.Status.Ziel_Geschwindigkeit;
   //--------------------------
         L     #IN_DW_Rampe_Pos;
         T     #Temp_IO_Status.Status.Ziel_Beschleunigung;
         L     #IN_DW_Rampe_Neg;
         T     #Temp_IO_Status.Status.Ziel_Verzoegerung;
   //--------------------------
   // Nachlaufzeit für Positionierung
         A     #Temp_IO_Status.Status.RT_dreht;
         L     S5T#500MS;
         SF    #IN_TM_Universal;
         A     #IN_TM_Universal;
         A     #Temp_FRG_Bewegung;
         =     #Temp_IO_Status.Ausgaenge_an_IPOS.DI_00_Start;
   ea_k: NOP   0;
END_REGION

REGION Network 17: Sollwerte an den Umrichter
         L     #Temp_IO_Status.Status.Ziel_Position;
         T     #Temp_IO_Status.Ausgaenge_an_IPOS.Zielposition;
   //--------------------------
         L     #Temp_IO_Status.Status.Ziel_Geschwindigkeit;
         T     #Temp_IO_Status.Ausgaenge_an_IPOS.Geschwindigkeit;
   //--------------------------
         L     #Temp_IO_Status.Status.Ziel_Beschleunigung;
         T     #Temp_IO_Status.Ausgaenge_an_IPOS.Positive_Rampe;
   //--------------------------
         L     #Temp_IO_Status.Status.Ziel_Verzoegerung;
         T     #Temp_IO_Status.Ausgaenge_an_IPOS.Negative_Rampe;
END_REGION

REGION Network 18: Kettenspanner anfordern
         O     #IN_BA_Hand;
         O     #IN_BA_Referenzieren;
         A(;
         O     #IN_T_Tippen_plus;
         O     #IN_T_Tippen_minus;
         );
         O     #IN_BA_Start_Taktbetrieb;
         O     #IN_BA_Taktbetrieb;
         =     #Temp_IO_Status.Status.Kettenspannung_noetig;
END_REGION

REGION Network 19: Freigaben an Umrichter
         L     S5T#2S;
         O     #Temp_IO_Status.Ausgaenge_an_IPOS.DI_00_Start;
         O     #Temp_IO_Status.Ausgaenge_an_IPOS.DI_01_T_plus;
         O     #Temp_IO_Status.Ausgaenge_an_IPOS.DI_02_T_minus;
         A     #Temp_FRG_Bewegung;
         SF    #IN_TM_Freigabe;
   //
         A     #IN_TM_Freigabe;
         =     #Temp_IO_Status.Ausgaenge_an_IPOS.Freigabe_Halt;
         =     #Temp_IO_Status.Ausgaenge_an_IPOS.Freigabe_Schnellstop;
   //
         A     #IN_HW_und_BA_ok;
         =     #OUT_FRG_Umrichter;
END_REGION

REGION Network 20: Lampenansteuerung
         A     #IN_BA_Hand;
         A     #Temp_IO_Status.Ausgaenge_an_IPOS.DI_01_T_plus;
         A     "Flag_01_000_Hertz";
         O     #Temp_IO_Status.Status.RT_in_Position;
         O     #IN_BA_Lampentest;
         =     #OUT_H_Tippen_plus;
   //
         A     #IN_BA_Hand;
         A     #Temp_IO_Status.Ausgaenge_an_IPOS.DI_02_T_minus;
         A     "Flag_01_000_Hertz";
         O     #Temp_IO_Status.Status.RT_in_Position;
         O     #IN_BA_Lampentest;
         =     #OUT_H_Tippen_minus;
   //
         A     #IN_IPOS_referenziert;
         =     #Temp_IO_Status.Status.IPOS_referenziert;
   //
         AN    #Temp_IO_Status.Status.IPOS_referenziert;
         R     #Temp_IO_Status.Status.RT_in_Position;
   //
         A     #IN_BA_Hand;
         A     #IN_BA_Referenzieren;
         A     #Temp_IO_Status.Ausgaenge_an_IPOS.DI_00_Start;
         A     "Flag_01_250_Hertz";
         O     #Temp_IO_Status.Status.IPOS_referenziert;
         O     #IN_BA_Lampentest;
         =     #OUT_H_Referenzpunkt;
END_REGION

REGION Network 21: Anfahrwarnungshupe ansteuern / Start verzögern
         A     #Temp_IO_Status.Ausgaenge_an_IPOS.Freigabe_Halt;
         L     #IN_Time_Anfahrwarnung;
         SD    #IN_TM_AnfahrWarnung;

   // Hupe ausgeben
         A     #Temp_IO_Status.Ausgaenge_an_IPOS.Freigabe_Halt;
         AN    #IN_TM_AnfahrWarnung;
         =     #OUT_H_AnfahrWarnung;

   // Starten wenn Warnung Ende
         A     #Temp_IO_Status.Ausgaenge_an_IPOS.Freigabe_Halt;
         A     #IN_TM_AnfahrWarnung;
         =     #Temp_IO_Status.Ausgaenge_an_IPOS.Freigabe_Halt;
END_REGION

REGION Network 22: Ausgänge an IPOS ausgeben
   // Um ein permanentes Beschreiben des Diagnosepuffers zu verhindern, werden die 
   // Peripheriebefehle übersprungen, sobald festgestellt wurde, daß der Teilnehmer 
   // ausgefallen ist.
         L     0;
         T     #Temp_Nullmerker;
   //
         AN    #IN_DP_ok;
         JC    paae;
   //
         CALL  DPWR_DAT
         ( LADDR   := #IN_EA_Adresse,
           RECORD  := #Temp_IO_Status.Ausgaenge_an_IPOS,
           RET_VAL := #ERROR_CODE
         );
   //
   paae: NOP   0;
END_REGION

REGION Network 23: Daten sichern
         CALL  BLKMOV
         ( SRCBLK  := #Temp_IO_Status,
           RET_VAL := #ERROR_CODE,
           DSTBLK  := #Anyzeiger
         );
   //
END_REGION
END_FUNCTION

FUNCTION "FC1043_RT_Segmentkennung" : Void   // FC1043, STL
TITLE = Segmentnummer in Station 1 ermitteln
{ S7_Optimized_Access := 'FALSE' }
AUTHOR : KT242
VERSION : 0.1
   VAR_INPUT
      IN_Segmentzahl : Int;   // Anzahl der vorhandenen Segmente
      IN_Muster_Last_SG_Stat_1 : DWord;   // Bitmuster der Segmentinis wenn das letzte Segment in der Station 1 steht
      IN_Segmentinis : DWord;   // Eingangswort mit den Eingängen der Segmentkennungen (Hardwareabschaltungen)
      IN_Segmente_Aufsteigend : Bool;   // Bedeutet die Drehrichtung eine aufsteigende Nummerierung der Segmente?
      IN_Anlage_in_Position : Bool;   // Die Anlage befindet sich in der vorgegebenen Position
      IN_Betriebsart_Automatik : Bool;   // Die Anlage befindet sich im Automatik- Betrieb
      IN_Reset_fault_Fkt : Bool;   // Signal zum quittieren der Störungen innerhalb der einzelnen Funktionsbausteine
   END_VAR
   VAR_IN_OUT
      IO_Status : "UDT_RT_Station_Nr";   // Speichern der Segmentkennungs- Zustände für das Programm
   END_VAR
   VAR_TEMP
      Temp_Schleifenzaehler : Int;   // Hilfswort für einen internen Schleifenzähler
      Temp_Seg_No_Stat_1 : Int;   // Hilfswort mit der Nummer des aktuellen Segmentes in der Position 1
      Temp_Testmuster : DWord;   // Hilfsdoppelwort für das Bitmuster zur Ermittelung des Segmentes in Position 1
      Temp_Segmentinis : DWord;   // Hilfsdoppelwort mit den aktuell benötigten Eingängen der Segmentinis
      Temp_Nummer_gleich : Bool;   // Hilfsmerker das die neue und die alte Nummer gleich sind
      Temp_Nummer_plus_1 : Bool;   // Hilfsmerker das die neue Nummer um 1 größer als die alte Nummer ist
      Temp_Nummer_minus_1 : Bool;   // Hilfsmerker das die neue Nummer um 1 kleiner als die alte Nummer ist
      Temp_Nummer_vorher_0 : Bool;   // Hilfsmerker das die alte Nummer 0 war
   END_VAR
BEGIN

REGION Network 1: Prüfen, zu welcher RT-Stellung das Eingangsmuster paßt
         L     #IN_Muster_Last_SG_Stat_1;
         CAD;
         T     #Temp_Testmuster;
   //
         A(;
         L     32;
         L     #IN_Segmentzahl;
         >=I;
         );
         A(;
         L     0;
         >I;
         );
         JC    arb;
         T     #IO_Status.Seg_No_Stat_1;
         T     #IO_Status.Bitmuster_Seg_No_Stat_1;
         BEU;
   // abhängig von der Anzahl der Segmente nicht benötigte Eingänge ausblenden
   arb:  NOP   0;
         L     #IN_Segmentinis;
         T     #Temp_Segmentinis;
   //
         L     #IN_Segmentzahl;
   m001: T     #Temp_Schleifenzaehler;
         L     #Temp_Segmentinis;
         CAD;
         L     #Temp_Testmuster;
         ==D;
         JC    nook;
         L     #Temp_Testmuster;
         SRD   1;  // neues Testmuster bilden
         T     #Temp_Testmuster;
         JZ    tneu;  // Sprung, wenn keine 1 geschoben
   //
         L     #IN_Segmentzahl;  // 1 an passender Stelle
         +     -1;  // einfügen, wenn eine 1
         L     DW#16#1;  // ausgeschoben wurde
         SLD;
         L     #Temp_Testmuster;
         OD;
         T     #Temp_Testmuster;
   //
   tneu: L     #Temp_Schleifenzaehler;
         LOOP  m001;
         T     #Temp_Schleifenzaehler;  // -> 0 falls Muster nicht gefunden
   //
   nook: L     #Temp_Schleifenzaehler;
         T     #Temp_Seg_No_Stat_1;
END_REGION

REGION Network 2: Störungsauswertung
   // Folgende Tests werden durchgeführt:
   // - bei Flanke auf eine temporäre Nummer <>0 wird geprüft, ob Nummer logisch paßt
   // - bei Rundtischstillstand wird geprüft, ob Nummer vorhanden ist
         A     #IN_Reset_fault_Fkt;
         R     #IO_Status.STG_Hardwareabschaltung;
         R     #IO_Status.STG_Nummer_unlogisch;
   //
   // Stationsnummer plus/minus feststellen
         A(;
         L     0;
         L     #IO_Status.Seg_No_Stat_1_alt;
         ==I;
         );
         A(;
         L     #Temp_Seg_No_Stat_1;
         <>I;
         T     #IO_Status.Seg_No_Stat_1_alt;
         );
         JC    test;
         JU    rpos;
   //
   test: O(;
         L     #IO_Status.Seg_No_Stat_1;
         +     1;
         L     #Temp_Seg_No_Stat_1;
         ==I;
         );
         O(;
         A(;
         L     #IO_Status.Seg_No_Stat_1;
         L     #IN_Segmentzahl;
         ==I;
         );
         A(;
         L     #Temp_Seg_No_Stat_1;
         L     1;
         ==I;
         );
         );
         =     #Temp_Nummer_plus_1;
   //
         O(;
         L     #Temp_Seg_No_Stat_1;
         +     1;
         L     #IO_Status.Seg_No_Stat_1;
         ==I;
         );
         O(;
         A(;
         L     #IO_Status.Seg_No_Stat_1;
         L     1;
         ==I;
         );
         A(;
         L     #Temp_Seg_No_Stat_1;
         L     #IN_Segmentzahl;
         ==I;
         );
         );
         =     #Temp_Nummer_minus_1;
   //
         L     #IO_Status.Seg_No_Stat_1;
         L     #Temp_Seg_No_Stat_1;
         ==I;
         =     #Temp_Nummer_gleich;
   //
         L     #IO_Status.Seg_No_Stat_1;
         L     0;
         ==I;
         =     #Temp_Nummer_vorher_0;
   //
         A(;
         AN    #Temp_Nummer_plus_1;
         AN    #Temp_Nummer_gleich;
         AN    #Temp_Nummer_minus_1;
         AN    #Temp_Nummer_vorher_0;
         O;
         A     #IN_Betriebsart_Automatik;
         A     #IN_Segmente_Aufsteigend;
         AN    #Temp_Nummer_plus_1;
         AN    #Temp_Nummer_vorher_0;
         O;
         A     #IN_Betriebsart_Automatik;
         AN    #IN_Segmente_Aufsteigend;
         AN    #Temp_Nummer_minus_1;
         AN    #Temp_Nummer_vorher_0;
         );
         A     #IN_Anlage_in_Position;
         S     #IO_Status.STG_Nummer_unlogisch;
   //
   rpos: A     #IN_Anlage_in_Position;
         A(;
         L     #Temp_Seg_No_Stat_1;
         L     0;
         ==I;
         );
         S     #IO_Status.STG_Hardwareabschaltung;
END_REGION

REGION Network 3: Ausgabe von Stationsnummer und Bitmuster
         AN    #IO_Status.STG_Hardwareabschaltung;
         AN    #IO_Status.STG_Nummer_unlogisch;
         JC    ausg;
         L     0;
         T     #IO_Status.Seg_No_Stat_1;
         JU    bits;
   ausg: NOP   0;
         O(;
         L     0;
         L     #Temp_Seg_No_Stat_1;
         ==I;
         );
         ON    #IN_Anlage_in_Position;
         JC    ende;
         T     #IO_Status.Seg_No_Stat_1;
   // Bitmuster bilden
   bits: L     0;
         L     #IO_Status.Seg_No_Stat_1;
         ==I;
         JC    tran;
         DEC   1;
         L     W#16#1;
         SLD;
   tran: T     #IO_Status.Bitmuster_Seg_No_Stat_1;
   ende: BE;
END_REGION
END_FUNCTION

FUNCTION "FC1044_Kettenspanner" : Void   // FC1044, STL
TITLE = Kettenspanner
{ S7_Optimized_Access := 'FALSE' }
AUTHOR : KT242